   1541: 'Carrier 24 CB02123 Tripped', class No Acknowledgement, trigger "DB302_HMI_Faults_Carrier24_Faults_0" bit 4
   1542: 'Carrier 24 AUX1 CB Tripped', class No Acknowledgement, trigger "DB302_HMI_Faults_Carrier24_Faults_0" bit 5
   1543: 'Carrier 24 AUX2 CB Tripped', class No Acknowledgement, trigger "DB302_HMI_Faults_Carrier24_Faults_0" bit 6
   1544: 'Carrier 24 PLC Not Communicating', class No Acknowledgement, trigger "DB302_HMI_Faults_Carrier24_Faults_0" bit 7
   1545: 'Carrier 24 Safe Input Card Fault', class No Acknowledgement, trigger "DB302_HMI_Faults_Carrier24_Faults_0" bit 8
   1546: 'Carrier 24 Safe Output Card Fault', class No Acknowledgement, trigger "DB302_HMI_Faults_Carrier24_Faults_0" bit 9
   1547: 'Carrier 24 Standard Input Card Fault', class No Acknowledgement, trigger "DB302_HMI_Faults_Carrier24_Faults_0" bit 10
   1548: 'Carrier 24 Standard Output Card Fault', class No Acknowledgement, trigger "DB302_HMI_Faults_Carrier24_Faults_0" bit 11
   1549: 'Carrier 24 Encoder Position Fault', class No Acknowledgement, trigger "DB302_HMI_Faults_Carrier24_Faults_0" bit 12
   1550: 'Carrier 24 Encoder Internal Error', class No Acknowledgement, trigger "DB302_HMI_Faults_Carrier24_Faults_0" bit 13
   1551: 'Carrier 24 Encoder Comm Fault', class No Acknowledgement, trigger "DB302_HMI_Faults_Carrier24_Faults_0" bit 14
   1552: 'Carrier 24 HMI Comm Fault', class No Acknowledgement, trigger "DB302_HMI_Faults_Carrier24_Faults_0" bit 15
   1553: 'Carrier 24 Crash Detection Fault', class No Acknowledgement, trigger "DB302_HMI_Faults_Carrier24_Faults_1" bit 0
   1554: 'Carrier 24 Carrier Number Invalid', class No Acknowledgement, trigger "DB302_HMI_Faults_Carrier24_Faults_1" bit 1
   1555: 'Carrier 24 Drive: PROFINET configuration error', class No Acknowledgement, trigger "DB302_HMI_Faults_Carrier24_Faults_1" bit 2
   1556: 'Carrier 24 Drive: Error internal communications', class No Acknowledgement, trigger "DB302_HMI_Faults_Carrier24_Faults_1" bit 3
   1557: 'Carrier 24 Drive: Motor overtemperature', class No Acknowledgement, trigger "DB302_HMI_Faults_Carrier24_Faults_1" bit 4
   1558: 'Carrier 24 Drive: Motor overcurrent', class No Acknowledgement, trigger "DB302_HMI_Faults_Carrier24_Faults_1" bit 5
   1559: 'Carrier 24 Drive: Infeed or power unit not ready', class No Acknowledgement, trigger "DB302_HMI_Faults_Carrier24_Faults_1" bit 6
   1560: 'Carrier 24 Drive: Short-circuit/ground fault detected', class No Acknowledgement, trigger "DB302_HMI_Faults_Carrier24_Faults_1" bit 7
   1561: 'Carrier 24 Drive: PROFINET Setpoint timeout', class No Acknowledgement, trigger "DB302_HMI_Faults_Carrier24_Faults_1" bit 8
   1562: 'Carrier 24 Power unit: Overcurrent', class No Acknowledgement, trigger "DB302_HMI_Faults_Carrier24_Faults_1" bit 9
   1563: 'Carrier 24 Power unit: DC link voltage overvoltage', class No Acknowledgement, trigger "DB302_HMI_Faults_Carrier24_Faults_1" bit 10
   1564: 'Carrier 24 Power unit: DC link voltage undervoltage', class No Acknowledgement, trigger "DB302_HMI_Faults_Carrier24_Faults_1" bit 11
   1565: 'Carrier 24 Power unit: Line phase failure in main circuit', class No Acknowledgement, trigger "DB302_HMI_Faults_Carrier24_Faults_1" bit 12
   1566: 'Carrier 24 Power unit: Phase failure motor cable', class No Acknowledgement, trigger "DB302_HMI_Faults_Carrier24_Faults_1" bit 13
   1567: 'Carrier 24 Power unit: Ground fault', class No Acknowledgement, trigger "DB302_HMI_Faults_Carrier24_Faults_1" bit 14
   1568: 'Spare_Fault_1568', class No Acknowledgement, trigger "DB302_HMI_Faults_Carrier24_Faults_1" bit 15
   1569: 'Carrier 24 Motion Off Fault', class No Acknowledgement, trigger "DB302_HMI_Faults_Carrier24_Faults_2" bit 0
   1570: 'Carrier 24 Motion On Fault', class No Acknowledgement, trigger "DB302_HMI_Faults_Carrier24_Faults_2" bit 1
   1571: 'Carrier 24 Spacing Fault', class No Acknowledgement, trigger "DB302_HMI_Faults_Carrier24_Faults_2" bit 2
   1572: 'Carrier 24 Duplicate Carrier Number Fault', class No Acknowledgement, trigger "DB302_HMI_Faults_Carrier24_Faults_2" bit 3
   1573: 'Spare_Fault_1573', class No Acknowledgement, trigger "DB302_HMI_Faults_Carrier24_Faults_2" bit 4
   1574: 'Spare_Fault_1574', class No Acknowledgement, trigger "DB302_HMI_Faults_Carrier24_Faults_2" bit 5
   1575: 'Spare_Fault_1575', class No Acknowledgement, trigger "DB302_HMI_Faults_Carrier24_Faults_2" bit 6
   1576: 'Spare_Fault_1576', class No Acknowledgement, trigger "DB302_HMI_Faults_Carrier24_Faults_2" bit 7
   1577: 'Spare_Fault_1577', class No Acknowledgement, trigger "DB302_HMI_Faults_Carrier24_Faults_2" bit 8
   1578: 'Spare_Fault_1578', class No Acknowledgement, trigger "DB302_HMI_Faults_Carrier24_Faults_2" bit 9
   1579: 'Spare_Fault_1579', class No Acknowledgement, trigger "DB302_HMI_Faults_Carrier24_Faults_2" bit 10
   1580: 'Spare_Fault_1580', class No Acknowledgement, trigger "DB302_HMI_Faults_Carrier24_Faults_2" bit 11
   1581: 'Spare_Fault_1581', class No Acknowledgement, trigger "DB302_HMI_Faults_Carrier24_Faults_2" bit 12
   1582: 'Spare_Fault_1582', class No Acknowledgement, trigger "DB302_HMI_Faults_Carrier24_Faults_2" bit 13
   1583: 'Spare_Fault_1583', class No Acknowledgement, trigger "DB302_HMI_Faults_Carrier24_Faults_2" bit 14
   1584: 'Spare_Fault_1584', class No Acknowledgement, trigger "DB302_HMI_Faults_Carrier24_Faults_2" bit 15
   1585: 'Spare_Fault_1585', class No Acknowledgement, trigger "DB302_HMI_Faults_Carrier24_Faults_3" bit 0
   1586: 'Spare_Fault_1586', class No Acknowledgement, trigger "DB302_HMI_Faults_Carrier24_Faults_3" bit 1
   1587: 'Spare_Fault_1587', class No Acknowledgement, trigger "DB302_HMI_Faults_Carrier24_Faults_3" bit 2
   1588: 'Spare_Fault_1588', class No Acknowledgement, trigger "DB302_HMI_Faults_Carrier24_Faults_3" bit 3
   1589: 'Spare_Fault_1589', class No Acknowledgement, trigger "DB302_HMI_Faults_Carrier24_Faults_3" bit 4
   1590: 'Spare_Fault_1590', class No Acknowledgement, trigger "DB302_HMI_Faults_Carrier24_Faults_3" bit 5
   1591: 'Spare_Fault_1591', class No Acknowledgement, trigger "DB302_HMI_Faults_Carrier24_Faults_3" bit 6
   1592: 'Spare_Fault_1592', class No Acknowledgement, trigger "DB302_HMI_Faults_Carrier24_Faults_3" bit 7
   1593: 'Spare_Fault_1593', class No Acknowledgement, trigger "DB302_HMI_Faults_Carrier24_Faults_3" bit 8
   1594: 'Spare_Fault_1594', class No Acknowledgement, trigger "DB302_HMI_Faults_Carrier24_Faults_3" bit 9
   1595: 'Spare_Fault_1595', class No Acknowledgement, trigger "DB302_HMI_Faults_Carrier24_Faults_3" bit 10
   1596: 'Spare_Fault_1596', class No Acknowledgement, trigger "DB302_HMI_Faults_Carrier24_Faults_3" bit 11
   1597: 'Spare_Fault_1597', class No Acknowledgement, trigger "DB302_HMI_Faults_Carrier24_Faults_3" bit 12
   1598: 'Spare_Fault_1598', class No Acknowledgement, trigger "DB302_HMI_Faults_Carrier24_Faults_3" bit 13
   1599: 'Spare_Fault_1599', class No Acknowledgement, trigger "DB302_HMI_Faults_Carrier24_Faults_3" bit 14
   1600: 'Spare_Fault_1600', class No Acknowledgement, trigger "DB302_HMI_Faults_Carrier24_Faults_3" bit 15
   1601: 'Carrier 25 Disconnect Open Power Fault DI11.0', class No Acknowledgement, trigger "DB302_HMI_Faults_Carrier25_Faults_0" bit 0
   1602: 'Carrier 25 Drive Profinet Comm Fault', class No Acknowledgement, trigger "DB302_HMI_Faults_Carrier25_Faults_0" bit 1
   1603: 'Carrier 25 Production Stop Not Reset', class No Acknowledgement, trigger "DB302_HMI_Faults_Carrier25_Faults_0" bit 2
   1604: 'Carrier 25 CB02122 Tripped', class No Acknowledgement, trigger "DB302_HMI_Faults_Carrier25_Faults_0" bit 3
   1605: 'Carrier 25 CB02123 Tripped', class No Acknowledgement, trigger "DB302_HMI_Faults_Carrier25_Faults_0" bit 4
   1606: 'Carrier 25 AUX1 CB Tripped', class No Acknowledgement, trigger "DB302_HMI_Faults_Carrier25_Faults_0" bit 5
   1607: 'Carrier 25 AUX2 CB Tripped', class No Acknowledgement, trigger "DB302_HMI_Faults_Carrier25_Faults_0" bit 6
   1608: 'Carrier 25 PLC Not Communicating', class No Acknowledgement, trigger "DB302_HMI_Faults_Carrier25_Faults_0" bit 7
   1609: 'Carrier 25 Safe Input Card Fault', class No Acknowledgement, trigger "DB302_HMI_Faults_Carrier25_Faults_0" bit 8
   1610: 'Carrier 25 Safe Output Card Fault', class No Acknowledgement, trigger "DB302_HMI_Faults_Carrier25_Faults_0" bit 9
   1611: 'Carrier 25 Standard Input Card Fault', class No Acknowledgement, trigger "DB302_HMI_Faults_Carrier25_Faults_0" bit 10
   1612: 'Carrier 25 Standard Output Card Fault', class No Acknowledgement, trigger "DB302_HMI_Faults_Carrier25_Faults_0" bit 11
   1613: 'Carrier 25 Encoder Position Fault', class No Acknowledgement, trigger "DB302_HMI_Faults_Carrier25_Faults_0" bit 12
   1614: 'Carrier 25 Encoder Internal Error', class No Acknowledgement, trigger "DB302_HMI_Faults_Carrier25_Faults_0" bit 13
   1615: 'Carrier 25 Encoder Comm Fault', class No Acknowledgement, trigger "DB302_HMI_Faults_Carrier25_Faults_0" bit 14
   1616: 'Carrier 25 HMI Comm Fault', class No Acknowledgement, trigger "DB302_HMI_Faults_Carrier25_Faults_0" bit 15
   1617: 'Carrier 25 Crash Detection Fault', class No Acknowledgement, trigger "DB302_HMI_Faults_Carrier25_Faults_1" bit 0
   1618: 'Carrier 25 Carrier Number Invalid', class No Acknowledgement, trigger "DB302_HMI_Faults_Carrier25_Faults_1" bit 1
   1619: 'Carrier 25 Drive: PROFINET configuration error', class No Acknowledgement, trigger "DB302_HMI_Faults_Carrier25_Faults_1" bit 2
   1620: 'Carrier 25 Drive: Error internal communications', class No Acknowledgement, trigger "DB302_HMI_Faults_Carrier25_Faults_1" bit 3
   1621: 'Carrier 25 Drive: Motor overtemperature', class No Acknowledgement, trigger "DB302_HMI_Faults_Carrier25_Faults_1" bit 4
   1622: 'Carrier 25 Drive: Motor overcurrent', class No Acknowledgement, trigger "DB302_HMI_Faults_Carrier25_Faults_1" bit 5
   1623: 'Carrier 25 Drive: Infeed or power unit not ready', class No Acknowledgement, trigger "DB302_HMI_Faults_Carrier25_Faults_1" bit 6
   1624: 'Carrier 25 Drive: Short-circuit/ground fault detected', class No Acknowledgement, trigger "DB302_HMI_Faults_Carrier25_Faults_1" bit 7
   1625: 'Carrier 25 Drive: PROFINET Setpoint timeout', class No Acknowledgement, trigger "DB302_HMI_Faults_Carrier25_Faults_1" bit 8
   1626: 'Carrier 25 Power unit: Overcurrent', class No Acknowledgement, trigger "DB302_HMI_Faults_Carrier25_Faults_1" bit 9
   1627: 'Carrier 25 Power unit: DC link voltage overvoltage', class No Acknowledgement, trigger "DB302_HMI_Faults_Carrier25_Faults_1" bit 10
   1628: 'Carrier 25 Power unit: DC link voltage undervoltage', class No Acknowledgement, trigger "DB302_HMI_Faults_Carrier25_Faults_1" bit 11
   1629: 'Carrier 25 Power unit: Line phase failure in main circuit', class No Acknowledgement, trigger "DB302_HMI_Faults_Carrier25_Faults_1" bit 12
   1630: 'Carrier 25 Power unit: Phase failure motor cable', class No Acknowledgement, trigger "DB302_HMI_Faults_Carrier25_Faults_1" bit 13
   1631: 'Carrier 25 Power unit: Ground fault', class No Acknowledgement, trigger "DB302_HMI_Faults_Carrier25_Faults_1" bit 14
   1632: 'Spare_Fault_1632', class No Acknowledgement, trigger "DB302_HMI_Faults_Carrier25_Faults_1" bit 15
   1633: 'Carrier 25 Motion Off Fault', class No Acknowledgement, trigger "DB302_HMI_Faults_Carrier25_Faults_2" bit 0
   1634: 'Carrier 25 Motion On Fault', class No Acknowledgement, trigger "DB302_HMI_Faults_Carrier25_Faults_2" bit 1
   1635: 'Carrier 25 Spacing Fault', class No Acknowledgement, trigger "DB302_HMI_Faults_Carrier25_Faults_2" bit 2
   1636: 'Carrier 25 Duplicate Carrier Number Fault', class No Acknowledgement, trigger "DB302_HMI_Faults_Carrier25_Faults_2" bit 3
   1637: 'Spare_Fault_1637', class No Acknowledgement, trigger "DB302_HMI_Faults_Carrier25_Faults_2" bit 4
   1638: 'Spare_Fault_1638', class No Acknowledgement, trigger "DB302_HMI_Faults_Carrier25_Faults_2" bit 5
   1639: 'Spare_Fault_1639', class No Acknowledgement, trigger "DB302_HMI_Faults_Carrier25_Faults_2" bit 6
   1640: 'Spare_Fault_1640', class No Acknowledgement, trigger "DB302_HMI_Faults_Carrier25_Faults_2" bit 7
   1641: 'Spare_Fault_1641', class No Acknowledgement, trigger "DB302_HMI_Faults_Carrier25_Faults_2" bit 8
   1642: 'Spare_Fault_1642', class No Acknowledgement, trigger "DB302_HMI_Faults_Carrier25_Faults_2" bit 9
   1643: 'Spare_Fault_1643', class No Acknowledgement, trigger "DB302_HMI_Faults_Carrier25_Faults_2" bit 10
   1644: 'Spare_Fault_1644', class No Acknowledgement, trigger "DB302_HMI_Faults_Carrier25_Faults_2" bit 11
   1645: 'Spare_Fault_1645', class No Acknowledgement, trigger "DB302_HMI_Faults_Carrier25_Faults_2" bit 12
   1646: 'Spare_Fault_1646', class No Acknowledgement, trigger "DB302_HMI_Faults_Carrier25_Faults_2" bit 13
   1647: 'Spare_Fault_1647', class No Acknowledgement, trigger "DB302_HMI_Faults_Carrier25_Faults_2" bit 14
   1648: 'Spare_Fault_1648', class No Acknowledgement, trigger "DB302_HMI_Faults_Carrier25_Faults_2" bit 15
   1649: 'Spare_Fault_1649', class No Acknowledgement, trigger "DB302_HMI_Faults_Carrier25_Faults_3" bit 0
   1650: 'Spare_Fault_1650', class No Acknowledgement, trigger "DB302_HMI_Faults_Carrier25_Faults_3" bit 1
   1651: 'Spare_Fault_1651', class No Acknowledgement, trigger "DB302_HMI_Faults_Carrier25_Faults_3" bit 2
   1652: 'Spare_Fault_1652', class No Acknowledgement, trigger "DB302_HMI_Faults_Carrier25_Faults_3" bit 3
   1653: 'Spare_Fault_1653', class No Acknowledgement, trigger "DB302_HMI_Faults_Carrier25_Faults_3" bit 4
   1654: 'Spare_Fault_1654', class No Acknowledgement, trigger "DB302_HMI_Faults_Carrier25_Faults_3" bit 5
   1655: 'Spare_Fault_1655', class No Acknowledgement, trigger "DB302_HMI_Faults_Carrier25_Faults_3" bit 6
   1656: 'Spare_Fault_1656', class No Acknowledgement, trigger "DB302_HMI_Faults_Carrier25_Faults_3" bit 7
   1657: 'Spare_Fault_1657', class No Acknowledgement, trigger "DB302_HMI_Faults_Carrier25_Faults_3" bit 8
   1658: 'Spare_Fault_1658', class No Acknowledgement, trigger "DB302_HMI_Faults_Carrier25_Faults_3" bit 9
   1659: 'Spare_Fault_1659', class No Acknowledgement, trigger "DB302_HMI_Faults_Carrier25_Faults_3" bit 10
   1660: 'Spare_Fault_1660', class No Acknowledgement, trigger "DB302_HMI_Faults_Carrier25_Faults_3" bit 11
   1661: 'Spare_Fault_1661', class No Acknowledgement, trigger "DB302_HMI_Faults_Carrier25_Faults_3" bit 12
   1662: 'Spare_Fault_1662', class No Acknowledgement, trigger "DB302_HMI_Faults_Carrier25_Faults_3" bit 13
   1663: 'Spare_Fault_1663', class No Acknowledgement, trigger "DB302_HMI_Faults_Carrier25_Faults_3" bit 14
   1664: 'Spare_Fault_1664', class No Acknowledgement, trigger "DB302_HMI_Faults_Carrier25_Faults_3" bit 15
   1665: 'Carrier 26 Disconnect Open Power Fault DI11.0', class No Acknowledgement, trigger "DB302_HMI_Faults_Carrier26_Faults_0" bit 0
   1666: 'Carrier 26 Drive Profinet Comm Fault', class No Acknowledgement, trigger "DB302_HMI_Faults_Carrier26_Faults_0" bit 1
   1667: 'Carrier 26 Production Stop Not Reset', class No Acknowledgement, trigger "DB302_HMI_Faults_Carrier26_Faults_0" bit 2
   1668: 'Carrier 26 CB02122 Tripped', class No Acknowledgement, trigger "DB302_HMI_Faults_Carrier26_Faults_0" bit 3
   1669: 'Carrier 26 CB02123 Tripped', class No Acknowledgement, trigger "DB302_HMI_Faults_Carrier26_Faults_0" bit 4
   1670: 'Carrier 26 AUX1 CB Tripped', class No Acknowledgement, trigger "DB302_HMI_Faults_Carrier26_Faults_0" bit 5
   1671: 'Carrier 26 AUX2 CB Tripped', class No Acknowledgement, trigger "DB302_HMI_Faults_Carrier26_Faults_0" bit 6
   1672: 'Carrier 26 PLC Not Communicating', class No Acknowledgement, trigger "DB302_HMI_Faults_Carrier26_Faults_0" bit 7
   1673: 'Carrier 26 Safe Input Card Fault', class No Acknowledgement, trigger "DB302_HMI_Faults_Carrier26_Faults_0" bit 8
   1674: 'Carrier 26 Safe Output Card Fault', class No Acknowledgement, trigger "DB302_HMI_Faults_Carrier26_Faults_0" bit 9
   1675: 'Carrier 26 Standard Input Card Fault', class No Acknowledgement, trigger "DB302_HMI_Faults_Carrier26_Faults_0" bit 10
   1676: 'Carrier 26 Standard Output Card Fault', class No Acknowledgement, trigger "DB302_HMI_Faults_Carrier26_Faults_0" bit 11
   1677: 'Carrier 26 Encoder Position Fault', class No Acknowledgement, trigger "DB302_HMI_Faults_Carrier26_Faults_0" bit 12
   1678: 'Carrier 26 Encoder Internal Error', class No Acknowledgement, trigger "DB302_HMI_Faults_Carrier26_Faults_0" bit 13
   1679: 'Carrier 26 Encoder Comm Fault', class No Acknowledgement, trigger "DB302_HMI_Faults_Carrier26_Faults_0" bit 14
   1680: 'Carrier 26 HMI Comm Fault', class No Acknowledgement, trigger "DB302_HMI_Faults_Carrier26_Faults_0" bit 15
   1681: 'Carrier 26 Crash Detection Fault', class No Acknowledgement, trigger "DB302_HMI_Faults_Carrier26_Faults_1" bit 0
   1682: 'Carrier 26 Carrier Number Invalid', class No Acknowledgement, trigger "DB302_HMI_Faults_Carrier26_Faults_1" bit 1
   1683: 'Carrier 26 Drive: PROFINET configuration error', class No Acknowledgement, trigger "DB302_HMI_Faults_Carrier26_Faults_1" bit 2
   1684: 'Carrier 26 Drive: Error internal communications', class No Acknowledgement, trigger "DB302_HMI_Faults_Carrier26_Faults_1" bit 3
   1685: 'Carrier 26 Drive: Motor overtemperature', class No Acknowledgement, trigger "DB302_HMI_Faults_Carrier26_Faults_1" bit 4
   1686: 'Carrier 26 Drive: Motor overcurrent', class No Acknowledgement, trigger "DB302_HMI_Faults_Carrier26_Faults_1" bit 5
   1687: 'Carrier 26 Drive: Infeed or power unit not ready', class No Acknowledgement, trigger "DB302_HMI_Faults_Carrier26_Faults_1" bit 6
   1688: 'Carrier 26 Drive: Short-circuit/ground fault detected', class No Acknowledgement, trigger "DB302_HMI_Faults_Carrier26_Faults_1" bit 7
   1689: 'Carrier 26 Drive: PROFINET Setpoint timeout', class No Acknowledgement, trigger "DB302_HMI_Faults_Carrier26_Faults_1" bit 8
   1690: 'Carrier 26 Power unit: Overcurrent', class No Acknowledgement, trigger "DB302_HMI_Faults_Carrier26_Faults_1" bit 9
   1691: 'Carrier 26 Power unit: DC link voltage overvoltage', class No Acknowledgement, trigger "DB302_HMI_Faults_Carrier26_Faults_1" bit 10
   1692: 'Carrier 26 Power unit: DC link voltage undervoltage', class No Acknowledgement, trigger "DB302_HMI_Faults_Carrier26_Faults_1" bit 11
   1693: 'Carrier 26 Power unit: Line phase failure in main circuit', class No Acknowledgement, trigger "DB302_HMI_Faults_Carrier26_Faults_1" bit 12
   1694: 'Carrier 26 Power unit: Phase failure motor cable', class No Acknowledgement, trigger "DB302_HMI_Faults_Carrier26_Faults_1" bit 13
   1695: 'Carrier 26 Power unit: Ground fault', class No Acknowledgement, trigger "DB302_HMI_Faults_Carrier26_Faults_1" bit 14
   1696: 'Spare_Fault_1696', class No Acknowledgement, trigger "DB302_HMI_Faults_Carrier26_Faults_1" bit 15
   1697: 'Carrier 26 Motion Off Fault', class No Acknowledgement, trigger "DB302_HMI_Faults_Carrier26_Faults_2" bit 0
   1698: 'Carrier 26 Motion On Fault', class No Acknowledgement, trigger "DB302_HMI_Faults_Carrier26_Faults_2" bit 1
   1699: 'Carrier 26 Spacing Fault', class No Acknowledgement, trigger "DB302_HMI_Faults_Carrier26_Faults_2" bit 2
   1700: 'Carrier 26 Duplicate Carrier Number Fault', class No Acknowledgement, trigger "DB302_HMI_Faults_Carrier26_Faults_2" bit 3
   1701: 'Spare_Fault_1701', class No Acknowledgement, trigger "DB302_HMI_Faults_Carrier26_Faults_2" bit 4
   1702: 'Spare_Fault_1702', class No Acknowledgement, trigger "DB302_HMI_Faults_Carrier26_Faults_2" bit 5
   1703: 'Spare_Fault_1703', class No Acknowledgement, trigger "DB302_HMI_Faults_Carrier26_Faults_2" bit 6
   1704: 'Spare_Fault_1704', class No Acknowledgement, trigger "DB302_HMI_Faults_Carrier26_Faults_2" bit 7
   1705: 'Spare_Fault_1705', class No Acknowledgement, trigger "DB302_HMI_Faults_Carrier26_Faults_2" bit 8
   1706: 'Spare_Fault_1706', class No Acknowledgement, trigger "DB302_HMI_Faults_Carrier26_Faults_2" bit 9
   1707: 'Spare_Fault_1707', class No Acknowledgement, trigger "DB302_HMI_Faults_Carrier26_Faults_2" bit 10
   1708: 'Spare_Fault_1708', class No Acknowledgement, trigger "DB302_HMI_Faults_Carrier26_Faults_2" bit 11
   1709: 'Spare_Fault_1709', class No Acknowledgement, trigger "DB302_HMI_Faults_Carrier26_Faults_2" bit 12
   1710: 'Spare_Fault_1710', class No Acknowledgement, trigger "DB302_HMI_Faults_Carrier26_Faults_2" bit 13
   1711: 'Spare_Fault_1711', class No Acknowledgement, trigger "DB302_HMI_Faults_Carrier26_Faults_2" bit 14
   1712: 'Spare_Fault_1712', class No Acknowledgement, trigger "DB302_HMI_Faults_Carrier26_Faults_2" bit 15
   1713: 'Spare_Fault_1713', class No Acknowledgement, trigger "DB302_HMI_Faults_Carrier26_Faults_3" bit 0
   1714: 'Spare_Fault_1714', class No Acknowledgement, trigger "DB302_HMI_Faults_Carrier26_Faults_3" bit 1
   1715: 'Spare_Fault_1715', class No Acknowledgement, trigger "DB302_HMI_Faults_Carrier26_Faults_3" bit 2
   1716: 'Spare_Fault_1716', class No Acknowledgement, trigger "DB302_HMI_Faults_Carrier26_Faults_3" bit 3
   1717: 'Spare_Fault_1717', class No Acknowledgement, trigger "DB302_HMI_Faults_Carrier26_Faults_3" bit 4
   1718: 'Spare_Fault_1718', class No Acknowledgement, trigger "DB302_HMI_Faults_Carrier26_Faults_3" bit 5
   1719: 'Spare_Fault_1719', class No Acknowledgement, trigger "DB302_HMI_Faults_Carrier26_Faults_3" bit 6
   1720: 'Spare_Fault_1720', class No Acknowledgement, trigger "DB302_HMI_Faults_Carrier26_Faults_3" bit 7
   1721: 'Spare_Fault_1721', class No Acknowledgement, trigger "DB302_HMI_Faults_Carrier26_Faults_3" bit 8
   1722: 'Spare_Fault_1722', class No Acknowledgement, trigger "DB302_HMI_Faults_Carrier26_Faults_3" bit 9
   1723: 'Spare_Fault_1723', class No Acknowledgement, trigger "DB302_HMI_Faults_Carrier26_Faults_3" bit 10
   1724: 'Spare_Fault_1724', class No Acknowledgement, trigger "DB302_HMI_Faults_Carrier26_Faults_3" bit 11
   1725: 'Spare_Fault_1725', class No Acknowledgement, trigger "DB302_HMI_Faults_Carrier26_Faults_3" bit 12
   1726: 'Spare_Fault_1726', class No Acknowledgement, trigger "DB302_HMI_Faults_Carrier26_Faults_3" bit 13
   1727: 'Spare_Fault_1727', class No Acknowledgement, trigger "DB302_HMI_Faults_Carrier26_Faults_3" bit 14
   1728: 'Spare_Fault_1728', class No Acknowledgement, trigger "DB302_HMI_Faults_Carrier26_Faults_3" bit 15
   1729: 'Carrier 27 Disconnect Open Power Fault DI11.0', class No Acknowledgement, trigger "DB302_HMI_Faults_Carrier27_Faults_0" bit 0
   1730: 'Carrier 27 Drive Profinet Comm Fault', class No Acknowledgement, trigger "DB302_HMI_Faults_Carrier27_Faults_0" bit 1
   1731: 'Carrier 27 Production Stop Not Reset', class No Acknowledgement, trigger "DB302_HMI_Faults_Carrier27_Faults_0" bit 2
   1732: 'Carrier 27 CB02122 Tripped', class No Acknowledgement, trigger "DB302_HMI_Faults_Carrier27_Faults_0" bit 3
   1733: 'Carrier 27 CB02123 Tripped', class No Acknowledgement, trigger "DB302_HMI_Faults_Carrier27_Faults_0" bit 4
   1734: 'Carrier 27 AUX1 CB Tripped', class No Acknowledgement, trigger "DB302_HMI_Faults_Carrier27_Faults_0" bit 5
   1735: 'Carrier 27 AUX2 CB Tripped', class No Acknowledgement, trigger "DB302_HMI_Faults_Carrier27_Faults_0" bit 6
   1736: 'Carrier 27 PLC Not Communicating', class No Acknowledgement, trigger "DB302_HMI_Faults_Carrier27_Faults_0" bit 7
   1737: 'Carrier 27 Safe Input Card Fault', class No Acknowledgement, trigger "DB302_HMI_Faults_Carrier27_Faults_0" bit 8
   1738: 'Carrier 27 Safe Output Card Fault', class No Acknowledgement, trigger "DB302_HMI_Faults_Carrier27_Faults_0" bit 9
   1739: 'Carrier 27 Standard Input Card Fault', class No Acknowledgement, trigger "DB302_HMI_Faults_Carrier27_Faults_0" bit 10
   1740: 'Carrier 27 Standard Output Card Fault', class No Acknowledgement, trigger "DB302_HMI_Faults_Carrier27_Faults_0" bit 11
   1741: 'Carrier 27 Encoder Position Fault', class No Acknowledgement, trigger "DB302_HMI_Faults_Carrier27_Faults_0" bit 12
   1742: 'Carrier 27 Encoder Internal Error', class No Acknowledgement, trigger "DB302_HMI_Faults_Carrier27_Faults_0" bit 13
   1743: 'Carrier 27 Encoder Comm Fault', class No Acknowledgement, trigger "DB302_HMI_Faults_Carrier27_Faults_0" bit 14
   1744: 'Carrier 27 HMI Comm Fault', class No Acknowledgement, trigger "DB302_HMI_Faults_Carrier27_Faults_0" bit 15
   1745: 'Carrier 27 Crash Detection Fault', class No Acknowledgement, trigger "DB302_HMI_Faults_Carrier27_Faults_1" bit 0
   1746: 'Carrier 27 Carrier Number Invalid', class No Acknowledgement, trigger "DB302_HMI_Faults_Carrier27_Faults_1" bit 1
   1747: 'Carrier 27 Drive: PROFINET configuration error', class No Acknowledgement, trigger "DB302_HMI_Faults_Carrier27_Faults_1" bit 2
   1748: 'Carrier 27 Drive: Error internal communications', class No Acknowledgement, trigger "DB302_HMI_Faults_Carrier27_Faults_1" bit 3
   1749: 'Carrier 27 Drive: Motor overtemperature', class No Acknowledgement, trigger "DB302_HMI_Faults_Carrier27_Faults_1" bit 4
   1750: 'Carrier 27 Drive: Motor overcurrent', class No Acknowledgement, trigger "DB302_HMI_Faults_Carrier27_Faults_1" bit 5
   1751: 'Carrier 27 Drive: Infeed or power unit not ready', class No Acknowledgement, trigger "DB302_HMI_Faults_Carrier27_Faults_1" bit 6
   1752: 'Carrier 27 Drive: Short-circuit/ground fault detected', class No Acknowledgement, trigger "DB302_HMI_Faults_Carrier27_Faults_1" bit 7
   1753: 'Carrier 27 Drive: PROFINET Setpoint timeout', class No Acknowledgement, trigger "DB302_HMI_Faults_Carrier27_Faults_1" bit 8
   1754: 'Carrier 27 Power unit: Overcurrent', class No Acknowledgement, trigger "DB302_HMI_Faults_Carrier27_Faults_1" bit 9
   1755: 'Carrier 27 Power unit: DC link voltage overvoltage', class No Acknowledgement, trigger "DB302_HMI_Faults_Carrier27_Faults_1" bit 10
   1756: 'Carrier 27 Power unit: DC link voltage undervoltage', class No Acknowledgement, trigger "DB302_HMI_Faults_Carrier27_Faults_1" bit 11
   1757: 'Carrier 27 Power unit: Line phase failure in main circuit', class No Acknowledgement, trigger "DB302_HMI_Faults_Carrier27_Faults_1" bit 12
   1758: 'Carrier 27 Power unit: Phase failure motor cable', class No Acknowledgement, trigger "DB302_HMI_Faults_Carrier27_Faults_1" bit 13
   1759: 'Carrier 27 Power unit: Ground fault', class No Acknowledgement, trigger "DB302_HMI_Faults_Carrier27_Faults_1" bit 14
   1760: 'Spare_Fault_1760', class No Acknowledgement, trigger "DB302_HMI_Faults_Carrier27_Faults_1" bit 15
   1761: 'Carrier 27 Motion Off Fault', class No Acknowledgement, trigger "DB302_HMI_Faults_Carrier27_Faults_2" bit 0
   1762: 'Carrier 27 Motion On Fault', class No Acknowledgement, trigger "DB302_HMI_Faults_Carrier27_Faults_2" bit 1
   1763: 'Carrier 27 Spacing Fault', class No Acknowledgement, trigger "DB302_HMI_Faults_Carrier27_Faults_2" bit 2
   1764: 'Carrier 27 Duplicate Carrier Number Fault', class No Acknowledgement, trigger "DB302_HMI_Faults_Carrier27_Faults_2" bit 3
   1765: 'Spare_Fault_1765', class No Acknowledgement, trigger "DB302_HMI_Faults_Carrier27_Faults_2" bit 4
   1766: 'Spare_Fault_1766', class No Acknowledgement, trigger "DB302_HMI_Faults_Carrier27_Faults_2" bit 5
   1767: 'Spare_Fault_1767', class No Acknowledgement, trigger "DB302_HMI_Faults_Carrier27_Faults_2" bit 6
   1768: 'Spare_Fault_1768', class No Acknowledgement, trigger "DB302_HMI_Faults_Carrier27_Faults_2" bit 7
   1769: 'Spare_Fault_1769', class No Acknowledgement, trigger "DB302_HMI_Faults_Carrier27_Faults_2" bit 8
   1770: 'Spare_Fault_1770', class No Acknowledgement, trigger "DB302_HMI_Faults_Carrier27_Faults_2" bit 9
   1771: 'Spare_Fault_1771', class No Acknowledgement, trigger "DB302_HMI_Faults_Carrier27_Faults_2" bit 10
   1772: 'Spare_Fault_1772', class No Acknowledgement, trigger "DB302_HMI_Faults_Carrier27_Faults_2" bit 11
   1773: 'Spare_Fault_1773', class No Acknowledgement, trigger "DB302_HMI_Faults_Carrier27_Faults_2" bit 12
   1774: 'Spare_Fault_1774', class No Acknowledgement, trigger "DB302_HMI_Faults_Carrier27_Faults_2" bit 13
   1775: 'Spare_Fault_1775', class No Acknowledgement, trigger "DB302_HMI_Faults_Carrier27_Faults_2" bit 14
   1776: 'Spare_Fault_1776', class No Acknowledgement, trigger "DB302_HMI_Faults_Carrier27_Faults_2" bit 15
   1777: 'Spare_Fault_1777', class No Acknowledgement, trigger "DB302_HMI_Faults_Carrier27_Faults_3" bit 0
   1778: 'Spare_Fault_1778', class No Acknowledgement, trigger "DB302_HMI_Faults_Carrier27_Faults_3" bit 1
   1779: 'Spare_Fault_1779', class No Acknowledgement, trigger "DB302_HMI_Faults_Carrier27_Faults_3" bit 2
   1780: 'Spare_Fault_1780', class No Acknowledgement, trigger "DB302_HMI_Faults_Carrier27_Faults_3" bit 3
   1781: 'Spare_Fault_1781', class No Acknowledgement, trigger "DB302_HMI_Faults_Carrier27_Faults_3" bit 4
   1782: 'Spare_Fault_1782', class No Acknowledgement, trigger "DB302_HMI_Faults_Carrier27_Faults_3" bit 5
   1783: 'Spare_Fault_1783', class No Acknowledgement, trigger "DB302_HMI_Faults_Carrier27_Faults_3" bit 6
   1784: 'Spare_Fault_1784', class No Acknowledgement, trigger "DB302_HMI_Faults_Carrier27_Faults_3" bit 7
   1785: 'Spare_Fault_1785', class No Acknowledgement, trigger "DB302_HMI_Faults_Carrier27_Faults_3" bit 8
   1786: 'Spare_Fault_1786', class No Acknowledgement, trigger "DB302_HMI_Faults_Carrier27_Faults_3" bit 9
   1787: 'Spare_Fault_1787', class No Acknowledgement, trigger "DB302_HMI_Faults_Carrier27_Faults_3" bit 10
   1788: 'Spare_Fault_1788', class No Acknowledgement, trigger "DB302_HMI_Faults_Carrier27_Faults_3" bit 11
   1789: 'Spare_Fault_1789', class No Acknowledgement, trigger "DB302_HMI_Faults_Carrier27_Faults_3" bit 12
   1790: 'Spare_Fault_1790', class No Acknowledgement, trigger "DB302_HMI_Faults_Carrier27_Faults_3" bit 13
   1791: 'Spare_Fault_1791', class No Acknowledgement, trigger "DB302_HMI_Faults_Carrier27_Faults_3" bit 14
   1792: 'Spare_Fault_1792', class No Acknowledgement, trigger "DB302_HMI_Faults_Carrier27_Faults_3" bit 15
   1793: 'Carrier 28 Disconnect Open Power Fault DI11.0', class No Acknowledgement, trigger "DB302_HMI_Faults_Carrier28_Faults_0" bit 0
   1794: 'Carrier 28 Drive Profinet Comm Fault', class No Acknowledgement, trigger "DB302_HMI_Faults_Carrier28_Faults_0" bit 1
   1795: 'Carrier 28 Production Stop Not Reset', class No Acknowledgement, trigger "DB302_HMI_Faults_Carrier28_Faults_0" bit 2
   1796: 'Carrier 28 CB02122 Tripped', class No Acknowledgement, trigger "DB302_HMI_Faults_Carrier28_Faults_0" bit 3
   1797: 'Carrier 28 CB02123 Tripped', class No Acknowledgement, trigger "DB302_HMI_Faults_Carrier28_Faults_0" bit 4
   1798: 'Carrier 28 AUX1 CB Tripped', class No Acknowledgement, trigger "DB302_HMI_Faults_Carrier28_Faults_0" bit 5
   1799: 'Carrier 28 AUX2 CB Tripped', class No Acknowledgement, trigger "DB302_HMI_Faults_Carrier28_Faults_0" bit 6
   1800: 'Carrier 28 PLC Not Communicating', class No Acknowledgement, trigger "DB302_HMI_Faults_Carrier28_Faults_0" bit 7
   1801: 'Carrier 28 Safe Input Card Fault', class No Acknowledgement, trigger "DB302_HMI_Faults_Carrier28_Faults_0" bit 8
   1802: 'Carrier 28 Safe Output Card Fault', class No Acknowledgement, trigger "DB302_HMI_Faults_Carrier28_Faults_0" bit 9
   1803: 'Carrier 28 Standard Input Card Fault', class No Acknowledgement, trigger "DB302_HMI_Faults_Carrier28_Faults_0" bit 10
   1804: 'Carrier 28 Standard Output Card Fault', class No Acknowledgement, trigger "DB302_HMI_Faults_Carrier28_Faults_0" bit 11
   1805: 'Carrier 28 Encoder Position Fault', class No Acknowledgement, trigger "DB302_HMI_Faults_Carrier28_Faults_0" bit 12
   1806: 'Carrier 28 Encoder Internal Error', class No Acknowledgement, trigger "DB302_HMI_Faults_Carrier28_Faults_0" bit 13
   1807: 'Carrier 28 Encoder Comm Fault', class No Acknowledgement, trigger "DB302_HMI_Faults_Carrier28_Faults_0" bit 14
   1808: 'Carrier 28 HMI Comm Fault', class No Acknowledgement, trigger "DB302_HMI_Faults_Carrier28_Faults_0" bit 15
   1809: 'Carrier 28 Crash Detection Fault', class No Acknowledgement, trigger "DB302_HMI_Faults_Carrier28_Faults_1" bit 0
   1810: 'Carrier 28 Carrier Number Invalid', class No Acknowledgement, trigger "DB302_HMI_Faults_Carrier28_Faults_1" bit 1
   1811: 'Carrier 28 Drive: PROFINET configuration error', class No Acknowledgement, trigger "DB302_HMI_Faults_Carrier28_Faults_1" bit 2
   1812: 'Carrier 28 Drive: Error internal communications', class No Acknowledgement, trigger "DB302_HMI_Faults_Carrier28_Faults_1" bit 3
   1813: 'Carrier 28 Drive: Motor overtemperature', class No Acknowledgement, trigger "DB302_HMI_Faults_Carrier28_Faults_1" bit 4
   1814: 'Carrier 28 Drive: Motor overcurrent', class No Acknowledgement, trigger "DB302_HMI_Faults_Carrier28_Faults_1" bit 5
   1815: 'Carrier 28 Drive: Infeed or power unit not ready', class No Acknowledgement, trigger "DB302_HMI_Faults_Carrier28_Faults_1" bit 6
   1816: 'Carrier 28 Drive: Short-circuit/ground fault detected', class No Acknowledgement, trigger "DB302_HMI_Faults_Carrier28_Faults_1" bit 7
   1817: 'Carrier 28 Drive: PROFINET Setpoint timeout', class No Acknowledgement, trigger "DB302_HMI_Faults_Carrier28_Faults_1" bit 8
   1818: 'Carrier 28 Power unit: Overcurrent', class No Acknowledgement, trigger "DB302_HMI_Faults_Carrier28_Faults_1" bit 9
   1819: 'Carrier 28 Power unit: DC link voltage overvoltage', class No Acknowledgement, trigger "DB302_HMI_Faults_Carrier28_Faults_1" bit 10
   1820: 'Carrier 28 Power unit: DC link voltage undervoltage', class No Acknowledgement, trigger "DB302_HMI_Faults_Carrier28_Faults_1" bit 11
   1821: 'Carrier 28 Power unit: Line phase failure in main circuit', class No Acknowledgement, trigger "DB302_HMI_Faults_Carrier28_Faults_1" bit 12
   1822: 'Carrier 28 Power unit: Phase failure motor cable', class No Acknowledgement, trigger "DB302_HMI_Faults_Carrier28_Faults_1" bit 13
   1823: 'Carrier 28 Power unit: Ground fault', class No Acknowledgement, trigger "DB302_HMI_Faults_Carrier28_Faults_1" bit 14
   1824: 'Spare_Fault_1824', class No Acknowledgement, trigger "DB302_HMI_Faults_Carrier28_Faults_1" bit 15
   1825: 'Carrier 28 Motion Off Fault', class No Acknowledgement, trigger "DB302_HMI_Faults_Carrier28_Faults_2" bit 0
   1826: 'Carrier 28 Motion On Fault', class No Acknowledgement, trigger "DB302_HMI_Faults_Carrier28_Faults_2" bit 1
   1827: 'Carrier 28 Spacing Fault', class No Acknowledgement, trigger "DB302_HMI_Faults_Carrier28_Faults_2" bit 2
   1828: 'Carrier 28 Duplicate Carrier Number Fault', class No Acknowledgement, trigger "DB302_HMI_Faults_Carrier28_Faults_2" bit 3
   1829: 'Spare_Fault_1829', class No Acknowledgement, trigger "DB302_HMI_Faults_Carrier28_Faults_2" bit 4
   1830: 'Spare_Fault_1830', class No Acknowledgement, trigger "DB302_HMI_Faults_Carrier28_Faults_2" bit 5
   1831: 'Spare_Fault_1831', class No Acknowledgement, trigger "DB302_HMI_Faults_Carrier28_Faults_2" bit 6
   1832: 'Spare_Fault_1832', class No Acknowledgement, trigger "DB302_HMI_Faults_Carrier28_Faults_2" bit 7
   1833: 'Spare_Fault_1833', class No Acknowledgement, trigger "DB302_HMI_Faults_Carrier28_Faults_2" bit 8
   1834: 'Spare_Fault_1834', class No Acknowledgement, trigger "DB302_HMI_Faults_Carrier28_Faults_2" bit 9
   1835: 'Spare_Fault_1835', class No Acknowledgement, trigger "DB302_HMI_Faults_Carrier28_Faults_2" bit 10
   1836: 'Spare_Fault_1836', class No Acknowledgement, trigger "DB302_HMI_Faults_Carrier28_Faults_2" bit 11
   1837: 'Spare_Fault_1837', class No Acknowledgement, trigger "DB302_HMI_Faults_Carrier28_Faults_2" bit 12
   1838: 'Spare_Fault_1838', class No Acknowledgement, trigger "DB302_HMI_Faults_Carrier28_Faults_2" bit 13
   1839: 'Spare_Fault_1839', class No Acknowledgement, trigger "DB302_HMI_Faults_Carrier28_Faults_2" bit 14
   1840: 'Spare_Fault_1840', class No Acknowledgement, trigger "DB302_HMI_Faults_Carrier28_Faults_2" bit 15
   1841: 'Spare_Fault_1841', class No Acknowledgement, trigger "DB302_HMI_Faults_Carrier28_Faults_3" bit 0
   1842: 'Spare_Fault_1842', class No Acknowledgement, trigger "DB302_HMI_Faults_Carrier28_Faults_3" bit 1
   1843: 'Spare_Fault_1843', class No Acknowledgement, trigger "DB302_HMI_Faults_Carrier28_Faults_3" bit 2
   1844: 'Spare_Fault_1844', class No Acknowledgement, trigger "DB302_HMI_Faults_Carrier28_Faults_3" bit 3
   1845: 'Spare_Fault_1845', class No Acknowledgement, trigger "DB302_HMI_Faults_Carrier28_Faults_3" bit 4
   1846: 'Spare_Fault_1846', class No Acknowledgement, trigger "DB302_HMI_Faults_Carrier28_Faults_3" bit 5
   1847: 'Spare_Fault_1847', class No Acknowledgement, trigger "DB302_HMI_Faults_Carrier28_Faults_3" bit 6
   1848: 'Spare_Fault_1848', class No Acknowledgement, trigger "DB302_HMI_Faults_Carrier28_Faults_3" bit 7
   1849: 'Spare_Fault_1849', class No Acknowledgement, trigger "DB302_HMI_Faults_Carrier28_Faults_3" bit 8
   1850: 'Spare_Fault_1850', class No Acknowledgement, trigger "DB302_HMI_Faults_Carrier28_Faults_3" bit 9
   1851: 'Spare_Fault_1851', class No Acknowledgement, trigger "DB302_HMI_Faults_Carrier28_Faults_3" bit 10
   1852: 'Spare_Fault_1852', class No Acknowledgement, trigger "DB302_HMI_Faults_Carrier28_Faults_3" bit 11
   1853: 'Spare_Fault_1853', class No Acknowledgement, trigger "DB302_HMI_Faults_Carrier28_Faults_3" bit 12
   1854: 'Spare_Fault_1854', class No Acknowledgement, trigger "DB302_HMI_Faults_Carrier28_Faults_3" bit 13
   1855: 'Spare_Fault_1855', class No Acknowledgement, trigger "DB302_HMI_Faults_Carrier28_Faults_3" bit 14
   1856: 'Spare_Fault_1856', class No Acknowledgement, trigger "DB302_HMI_Faults_Carrier28_Faults_3" bit 15
   1857: 'Carrier 29 Disconnect Open Power Fault DI11.0', class No Acknowledgement, trigger "DB302_HMI_Faults_Carrier29_Faults_0" bit 0
   1858: 'Carrier 29 Drive Profinet Comm Fault', class No Acknowledgement, trigger "DB302_HMI_Faults_Carrier29_Faults_0" bit 1
   1859: 'Carrier 29 Production Stop Not Reset', class No Acknowledgement, trigger "DB302_HMI_Faults_Carrier29_Faults_0" bit 2
   1860: 'Carrier 29 CB02122 Tripped', class No Acknowledgement, trigger "DB302_HMI_Faults_Carrier29_Faults_0" bit 3
   1861: 'Carrier 29 CB02123 Tripped', class No Acknowledgement, trigger "DB302_HMI_Faults_Carrier29_Faults_0" bit 4
   1862: 'Carrier 29 AUX1 CB Tripped', class No Acknowledgement, trigger "DB302_HMI_Faults_Carrier29_Faults_0" bit 5
   1863: 'Carrier 29 AUX2 CB Tripped', class No Acknowledgement, trigger "DB302_HMI_Faults_Carrier29_Faults_0" bit 6
   1864: 'Carrier 29 PLC Not Communicating', class No Acknowledgement, trigger "DB302_HMI_Faults_Carrier29_Faults_0" bit 7
   1865: 'Carrier 29 Safe Input Card Fault', class No Acknowledgement, trigger "DB302_HMI_Faults_Carrier29_Faults_0" bit 8
   1866: 'Carrier 29 Safe Output Card Fault', class No Acknowledgement, trigger "DB302_HMI_Faults_Carrier29_Faults_0" bit 9
   1867: 'Carrier 29 Standard Input Card Fault', class No Acknowledgement, trigger "DB302_HMI_Faults_Carrier29_Faults_0" bit 10
   1868: 'Carrier 29 Standard Output Card Fault', class No Acknowledgement, trigger "DB302_HMI_Faults_Carrier29_Faults_0" bit 11
   1869: 'Carrier 29 Encoder Position Fault', class No Acknowledgement, trigger "DB302_HMI_Faults_Carrier29_Faults_0" bit 12
   1870: 'Carrier 29 Encoder Internal Error', class No Acknowledgement, trigger "DB302_HMI_Faults_Carrier29_Faults_0" bit 13
   1871: 'Carrier 29 Encoder Comm Fault', class No Acknowledgement, trigger "DB302_HMI_Faults_Carrier29_Faults_0" bit 14
   1872: 'Carrier 29 HMI Comm Fault', class No Acknowledgement, trigger "DB302_HMI_Faults_Carrier29_Faults_0" bit 15
   1873: 'Carrier 29 Crash Detection Fault', class No Acknowledgement, trigger "DB302_HMI_Faults_Carrier29_Faults_1" bit 0
   1874: 'Carrier 29 Carrier Number Invalid', class No Acknowledgement, trigger "DB302_HMI_Faults_Carrier29_Faults_1" bit 1
   1875: 'Carrier 29 Drive: PROFINET configuration error', class No Acknowledgement, trigger "DB302_HMI_Faults_Carrier29_Faults_1" bit 2
   1876: 'Carrier 29 Drive: Error internal communications', class No Acknowledgement, trigger "DB302_HMI_Faults_Carrier29_Faults_1" bit 3
   1877: 'Carrier 29 Drive: Motor overtemperature', class No Acknowledgement, trigger "DB302_HMI_Faults_Carrier29_Faults_1" bit 4
   1878: 'Carrier 29 Drive: Motor overcurrent', class No Acknowledgement, trigger "DB302_HMI_Faults_Carrier29_Faults_1" bit 5
   1879: 'Carrier 29 Drive: Infeed or power unit not ready', class No Acknowledgement, trigger "DB302_HMI_Faults_Carrier29_Faults_1" bit 6
   1880: 'Carrier 29 Drive: Short-circuit/ground fault detected', class No Acknowledgement, trigger "DB302_HMI_Faults_Carrier29_Faults_1" bit 7
   1881: 'Carrier 29 Drive: PROFINET Setpoint timeout', class No Acknowledgement, trigger "DB302_HMI_Faults_Carrier29_Faults_1" bit 8
   1882: 'Carrier 29 Power unit: Overcurrent', class No Acknowledgement, trigger "DB302_HMI_Faults_Carrier29_Faults_1" bit 9
   1883: 'Carrier 29 Power unit: DC link voltage overvoltage', class No Acknowledgement, trigger "DB302_HMI_Faults_Carrier29_Faults_1" bit 10
   1884: 'Carrier 29 Power unit: DC link voltage undervoltage', class No Acknowledgement, trigger "DB302_HMI_Faults_Carrier29_Faults_1" bit 11
   1885: 'Carrier 29 Power unit: Line phase failure in main circuit', class No Acknowledgement, trigger "DB302_HMI_Faults_Carrier29_Faults_1" bit 12
   1886: 'Carrier 29 Power unit: Phase failure motor cable', class No Acknowledgement, trigger "DB302_HMI_Faults_Carrier29_Faults_1" bit 13
   1887: 'Carrier 29 Power unit: Ground fault', class No Acknowledgement, trigger "DB302_HMI_Faults_Carrier29_Faults_1" bit 14
   1888: 'Spare_Fault_1888', class No Acknowledgement, trigger "DB302_HMI_Faults_Carrier29_Faults_1" bit 15
   1889: 'Carrier 29 Motion Off Fault', class No Acknowledgement, trigger "DB302_HMI_Faults_Carrier29_Faults_2" bit 0
   1890: 'Carrier 29 Motion On Fault', class No Acknowledgement, trigger "DB302_HMI_Faults_Carrier29_Faults_2" bit 1
   1891: 'Carrier 29 Spacing Fault', class No Acknowledgement, trigger "DB302_HMI_Faults_Carrier29_Faults_2" bit 2
   1892: 'Carrier 29 Duplicate Carrier Number Fault', class No Acknowledgement, trigger "DB302_HMI_Faults_Carrier29_Faults_2" bit 3
   1893: 'Spare_Fault_1893', class No Acknowledgement, trigger "DB302_HMI_Faults_Carrier29_Faults_2" bit 4
   1894: 'Spare_Fault_1894', class No Acknowledgement, trigger "DB302_HMI_Faults_Carrier29_Faults_2" bit 5
   1895: 'Spare_Fault_1895', class No Acknowledgement, trigger "DB302_HMI_Faults_Carrier29_Faults_2" bit 6
   1896: 'Spare_Fault_1896', class No Acknowledgement, trigger "DB302_HMI_Faults_Carrier29_Faults_2" bit 7
   1897: 'Spare_Fault_1897', class No Acknowledgement, trigger "DB302_HMI_Faults_Carrier29_Faults_2" bit 8
   1898: 'Spare_Fault_1898', class No Acknowledgement, trigger "DB302_HMI_Faults_Carrier29_Faults_2" bit 9
   1899: 'Spare_Fault_1899', class No Acknowledgement, trigger "DB302_HMI_Faults_Carrier29_Faults_2" bit 10
   1900: 'Spare_Fault_1900', class No Acknowledgement, trigger "DB302_HMI_Faults_Carrier29_Faults_2" bit 11
   1901: 'Spare_Fault_1901', class No Acknowledgement, trigger "DB302_HMI_Faults_Carrier29_Faults_2" bit 12
   1902: 'Spare_Fault_1902', class No Acknowledgement, trigger "DB302_HMI_Faults_Carrier29_Faults_2" bit 13
   1903: 'Spare_Fault_1903', class No Acknowledgement, trigger "DB302_HMI_Faults_Carrier29_Faults_2" bit 14
   1904: 'Spare_Fault_1904', class No Acknowledgement, trigger "DB302_HMI_Faults_Carrier29_Faults_2" bit 15
   1905: 'Spare_Fault_1905', class No Acknowledgement, trigger "DB302_HMI_Faults_Carrier29_Faults_3" bit 0
   1906: 'Spare_Fault_1906', class No Acknowledgement, trigger "DB302_HMI_Faults_Carrier29_Faults_3" bit 1
   1907: 'Spare_Fault_1907', class No Acknowledgement, trigger "DB302_HMI_Faults_Carrier29_Faults_3" bit 2
   1908: 'Spare_Fault_1908', class No Acknowledgement, trigger "DB302_HMI_Faults_Carrier29_Faults_3" bit 3
   1909: 'Spare_Fault_1909', class No Acknowledgement, trigger "DB302_HMI_Faults_Carrier29_Faults_3" bit 4
   1910: 'Spare_Fault_1910', class No Acknowledgement, trigger "DB302_HMI_Faults_Carrier29_Faults_3" bit 5
   1911: 'Spare_Fault_1911', class No Acknowledgement, trigger "DB302_HMI_Faults_Carrier29_Faults_3" bit 6
   1912: 'Spare_Fault_1912', class No Acknowledgement, trigger "DB302_HMI_Faults_Carrier29_Faults_3" bit 7
   1913: 'Spare_Fault_1913', class No Acknowledgement, trigger "DB302_HMI_Faults_Carrier29_Faults_3" bit 8
   1914: 'Spare_Fault_1914', class No Acknowledgement, trigger "DB302_HMI_Faults_Carrier29_Faults_3" bit 9
   1915: 'Spare_Fault_1915', class No Acknowledgement, trigger "DB302_HMI_Faults_Carrier29_Faults_3" bit 10
   1916: 'Spare_Fault_1916', class No Acknowledgement, trigger "DB302_HMI_Faults_Carrier29_Faults_3" bit 11
   1917: 'Spare_Fault_1917', class No Acknowledgement, trigger "DB302_HMI_Faults_Carrier29_Faults_3" bit 12
   1918: 'Spare_Fault_1918', class No Acknowledgement, trigger "DB302_HMI_Faults_Carrier29_Faults_3" bit 13
   1919: 'Spare_Fault_1919', class No Acknowledgement, trigger "DB302_HMI_Faults_Carrier29_Faults_3" bit 14
   1920: 'Spare_Fault_1920', class No Acknowledgement, trigger "DB302_HMI_Faults_Carrier29_Faults_3" bit 15
   1921: 'Carrier 30 Disconnect Open Power Fault DI11.0', class No Acknowledgement, trigger "DB302_HMI_Faults_Carrier30_Faults_0" bit 0
   1922: 'Carrier 30 Drive Profinet Comm Fault', class No Acknowledgement, trigger "DB302_HMI_Faults_Carrier30_Faults_0" bit 1
   1923: 'Carrier 30 Production Stop Not Reset', class No Acknowledgement, trigger "DB302_HMI_Faults_Carrier30_Faults_0" bit 2
   1924: 'Carrier 30 CB02122 Tripped', class No Acknowledgement, trigger "DB302_HMI_Faults_Carrier30_Faults_0" bit 3
   1925: 'Carrier 30 CB02123 Tripped', class No Acknowledgement, trigger "DB302_HMI_Faults_Carrier30_Faults_0" bit 4
   1926: 'Carrier 30 AUX1 CB Tripped', class No Acknowledgement, trigger "DB302_HMI_Faults_Carrier30_Faults_0" bit 5
   1927: 'Carrier 30 AUX2 CB Tripped', class No Acknowledgement, trigger "DB302_HMI_Faults_Carrier30_Faults_0" bit 6
   1928: 'Carrier 30 PLC Not Communicating', class No Acknowledgement, trigger "DB302_HMI_Faults_Carrier30_Faults_0" bit 7
   1929: 'Carrier 30 Safe Input Card Fault', class No Acknowledgement, trigger "DB302_HMI_Faults_Carrier30_Faults_0" bit 8
   1930: 'Carrier 30 Safe Output Card Fault', class No Acknowledgement, trigger "DB302_HMI_Faults_Carrier30_Faults_0" bit 9
   1931: 'Carrier 30 Standard Input Card Fault', class No Acknowledgement, trigger "DB302_HMI_Faults_Carrier30_Faults_0" bit 10
   1932: 'Carrier 30 Standard Output Card Fault', class No Acknowledgement, trigger "DB302_HMI_Faults_Carrier30_Faults_0" bit 11
   1933: 'Carrier 30 Encoder Position Fault', class No Acknowledgement, trigger "DB302_HMI_Faults_Carrier30_Faults_0" bit 12
   1934: 'Carrier 30 Encoder Internal Error', class No Acknowledgement, trigger "DB302_HMI_Faults_Carrier30_Faults_0" bit 13
   1935: 'Carrier 30 Encoder Comm Fault', class No Acknowledgement, trigger "DB302_HMI_Faults_Carrier30_Faults_0" bit 14
   1936: 'Carrier 30 HMI Comm Fault', class No Acknowledgement, trigger "DB302_HMI_Faults_Carrier30_Faults_0" bit 15
   1937: 'Carrier 30 Crash Detection Fault', class No Acknowledgement, trigger "DB302_HMI_Faults_Carrier30_Faults_1" bit 0
   1938: 'Carrier 30 Carrier Number Invalid', class No Acknowledgement, trigger "DB302_HMI_Faults_Carrier30_Faults_1" bit 1
   1939: 'Carrier 30 Drive: PROFINET configuration error', class No Acknowledgement, trigger "DB302_HMI_Faults_Carrier30_Faults_1" bit 2
   1940: 'Carrier 30 Drive: Error internal communications', class No Acknowledgement, trigger "DB302_HMI_Faults_Carrier30_Faults_1" bit 3
   1941: 'Carrier 30 Drive: Motor overtemperature', class No Acknowledgement, trigger "DB302_HMI_Faults_Carrier30_Faults_1" bit 4
   1942: 'Carrier 30 Drive: Motor overcurrent', class No Acknowledgement, trigger "DB302_HMI_Faults_Carrier30_Faults_1" bit 5
   1943: 'Carrier 30 Drive: Infeed or power unit not ready', class No Acknowledgement, trigger "DB302_HMI_Faults_Carrier30_Faults_1" bit 6
   1944: 'Carrier 30 Drive: Short-circuit/ground fault detected', class No Acknowledgement, trigger "DB302_HMI_Faults_Carrier30_Faults_1" bit 7
   1945: 'Carrier 30 Drive: PROFINET Setpoint timeout', class No Acknowledgement, trigger "DB302_HMI_Faults_Carrier30_Faults_1" bit 8
   1946: 'Carrier 30 Power unit: Overcurrent', class No Acknowledgement, trigger "DB302_HMI_Faults_Carrier30_Faults_1" bit 9
   1947: 'Carrier 30 Power unit: DC link voltage overvoltage', class No Acknowledgement, trigger "DB302_HMI_Faults_Carrier30_Faults_1" bit 10
   1948: 'Carrier 30 Power unit: DC link voltage undervoltage', class No Acknowledgement, trigger "DB302_HMI_Faults_Carrier30_Faults_1" bit 11
   1949: 'Carrier 30 Power unit: Line phase failure in main circuit', class No Acknowledgement, trigger "DB302_HMI_Faults_Carrier30_Faults_1" bit 12
   1950: 'Carrier 30 Power unit: Phase failure motor cable', class No Acknowledgement, trigger "DB302_HMI_Faults_Carrier30_Faults_1" bit 13
   1951: 'Carrier 30 Power unit: Ground fault', class No Acknowledgement, trigger "DB302_HMI_Faults_Carrier30_Faults_1" bit 14
   1952: 'Spare_Fault_1952', class No Acknowledgement, trigger "DB302_HMI_Faults_Carrier30_Faults_1" bit 15
   1953: 'Carrier 30 Motion Off Fault', class No Acknowledgement, trigger "DB302_HMI_Faults_Carrier30_Faults_2" bit 0
   1954: 'Carrier 30 Motion On Fault', class No Acknowledgement, trigger "DB302_HMI_Faults_Carrier30_Faults_2" bit 1
   1955: 'Carrier 30 Spacing Fault', class No Acknowledgement, trigger "DB302_HMI_Faults_Carrier30_Faults_2" bit 2
   1956: 'Carrier 30 Duplicate Carrier Number Fault', class No Acknowledgement, trigger "DB302_HMI_Faults_Carrier30_Faults_2" bit 3
   1957: 'Spare_Fault_1957', class No Acknowledgement, trigger "DB302_HMI_Faults_Carrier30_Faults_2" bit 4
   1958: 'Spare_Fault_1958', class No Acknowledgement, trigger "DB302_HMI_Faults_Carrier30_Faults_2" bit 5
   1959: 'Spare_Fault_1959', class No Acknowledgement, trigger "DB302_HMI_Faults_Carrier30_Faults_2" bit 6